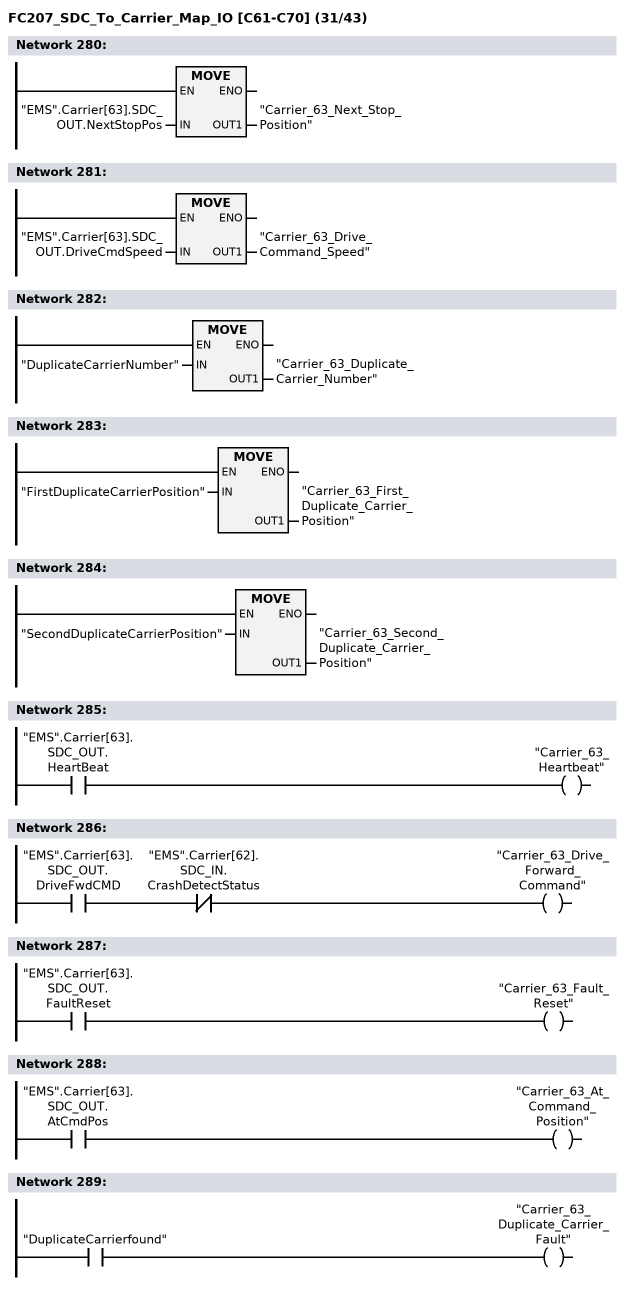
   RUNG wire#powerrail
      Move(in := "EMS".Carrier[63].SDC_OUT.NextStopPos, out1 => "Carrier_63_Next_Stop_Position")
   END_RUNG
   // the same network as SCL:
   "Carrier_63_Next_Stop_Position" := "EMS".Carrier[63].SDC_OUT.NextStopPos;
END_REGION

REGION Network 281
   RUNG wire#powerrail
      Move(in := "EMS".Carrier[63].SDC_OUT.DriveCmdSpeed, out1 => "Carrier_63_Drive_Command_Speed")
   END_RUNG
   // the same network as SCL:
   "Carrier_63_Drive_Command_Speed" := "EMS".Carrier[63].SDC_OUT.DriveCmdSpeed;
END_REGION

REGION Network 282
   RUNG wire#powerrail
      Move(in := "DuplicateCarrierNumber", out1 => "Carrier_63_Duplicate_Carrier_Number")
   END_RUNG
   // the same network as SCL:
   "Carrier_63_Duplicate_Carrier_Number" := "DuplicateCarrierNumber";
END_REGION

REGION Network 283
   RUNG wire#powerrail
      Move(in := "FirstDuplicateCarrierPosition", out1 => "Carrier_63_First_Duplicate_Carrier_Position")
   END_RUNG
   // the same network as SCL:
   "Carrier_63_First_Duplicate_Carrier_Position" := "FirstDuplicateCarrierPosition";
END_REGION

REGION Network 284
   RUNG wire#powerrail
      Move(in := "SecondDuplicateCarrierPosition", out1 => "Carrier_63_Second_Duplicate_Carrier_Position")
   END_RUNG
   // the same network as SCL:
   "Carrier_63_Second_Duplicate_Carrier_Position" := "SecondDuplicateCarrierPosition";
END_REGION

REGION Network 285
   RUNG wire#powerrail
      Contact( "EMS".Carrier[63].SDC_OUT.HeartBeat )
      Coil( "Carrier_63_Heartbeat" )
   END_RUNG
   // the same network as SCL:
   "Carrier_63_Heartbeat" := "EMS".Carrier[63].SDC_OUT.HeartBeat;
END_REGION

REGION Network 286
   RUNG wire#powerrail
      Contact( "EMS".Carrier[63].SDC_OUT.DriveFwdCMD )
      I_Contact( "EMS".Carrier[62].SDC_IN.CrashDetectStatus )
      Coil( "Carrier_63_Drive_Forward_Command" )
   END_RUNG
   // the same network as SCL:
   "Carrier_63_Drive_Forward_Command" := "EMS".Carrier[63].SDC_OUT.DriveFwdCMD AND NOT "EMS".Carrier[62].SDC_IN.CrashDetectStatus;
END_REGION

REGION Network 287
   RUNG wire#powerrail
      Contact( "EMS".Carrier[63].SDC_OUT.FaultReset )
      Coil( "Carrier_63_Fault_Reset" )
   END_RUNG
   // the same network as SCL:
   "Carrier_63_Fault_Reset" := "EMS".Carrier[63].SDC_OUT.FaultReset;
END_REGION

REGION Network 288
   RUNG wire#powerrail
      Contact( "EMS".Carrier[63].SDC_OUT.AtCmdPos )
      Coil( "Carrier_63_At_Command_Position" )
   END_RUNG
   // the same network as SCL:
   "Carrier_63_At_Command_Position" := "EMS".Carrier[63].SDC_OUT.AtCmdPos;
END_REGION

REGION Network 289
   RUNG wire#powerrail
      Contact( "DuplicateCarrierfound" )
      Coil( "Carrier_63_Duplicate_Carrier_Fault" )
   END_RUNG
   // the same network as SCL:
   "Carrier_63_Duplicate_Carrier_Fault" := "DuplicateCarrierfound";
END_REGION

REGION Network 290
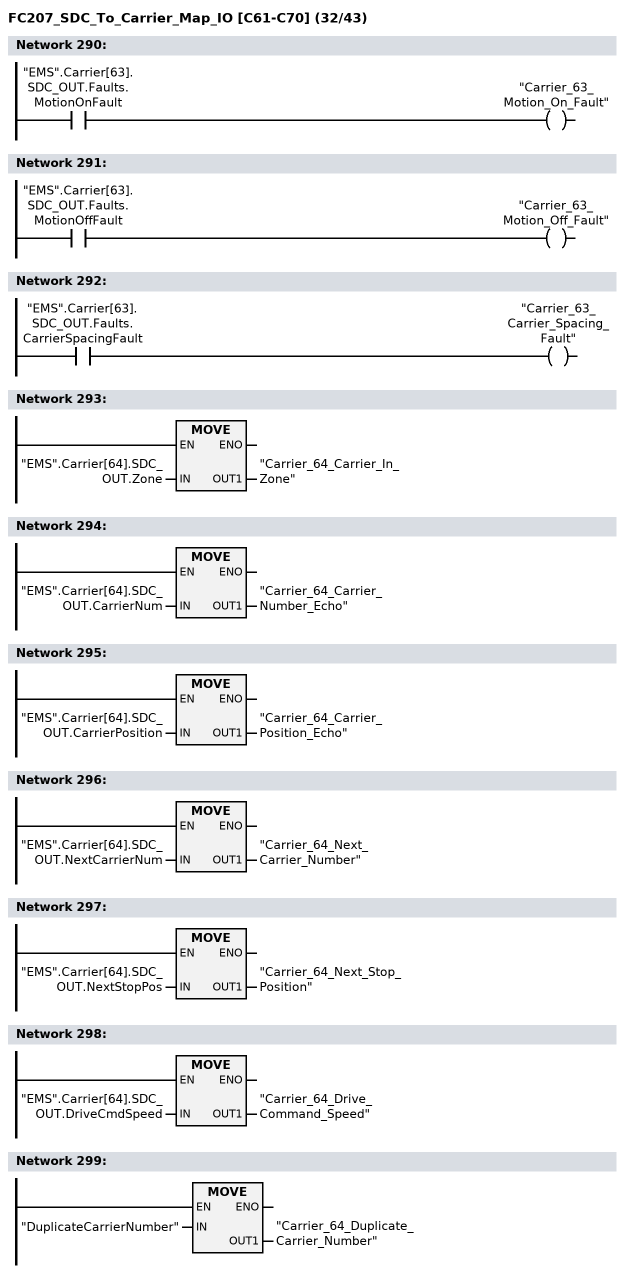
   RUNG wire#powerrail
      Contact( "EMS".Carrier[63].SDC_OUT.Faults.MotionOnFault )
      Coil( "Carrier_63_Motion_On_Fault" )
   END_RUNG
   // the same network as SCL:
   "Carrier_63_Motion_On_Fault" := "EMS".Carrier[63].SDC_OUT.Faults.MotionOnFault;
END_REGION

REGION Network 291
   RUNG wire#powerrail
      Contact( "EMS".Carrier[63].SDC_OUT.Faults.MotionOffFault )
      Coil( "Carrier_63_Motion_Off_Fault" )
   END_RUNG
   // the same network as SCL:
   "Carrier_63_Motion_Off_Fault" := "EMS".Carrier[63].SDC_OUT.Faults.MotionOffFault;
END_REGION

REGION Network 292
   RUNG wire#powerrail
      Contact( "EMS".Carrier[63].SDC_OUT.Faults.CarrierSpacingFault )
      Coil( "Carrier_63_Carrier_Spacing_Fault" )
   END_RUNG
   // the same network as SCL:
   "Carrier_63_Carrier_Spacing_Fault" := "EMS".Carrier[63].SDC_OUT.Faults.CarrierSpacingFault;
END_REGION

REGION Network 293
   RUNG wire#powerrail
      Move(in := "EMS".Carrier[64].SDC_OUT.Zone, out1 => "Carrier_64_Carrier_In_Zone")
   END_RUNG
   // the same network as SCL:
   "Carrier_64_Carrier_In_Zone" := "EMS".Carrier[64].SDC_OUT.Zone;
END_REGION

REGION Network 294
   RUNG wire#powerrail
      Move(in := "EMS".Carrier[64].SDC_OUT.CarrierNum, out1 => "Carrier_64_Carrier_Number_Echo")
   END_RUNG
   // the same network as SCL:
   "Carrier_64_Carrier_Number_Echo" := "EMS".Carrier[64].SDC_OUT.CarrierNum;
END_REGION

REGION Network 295
   RUNG wire#powerrail
      Move(in := "EMS".Carrier[64].SDC_OUT.CarrierPosition, out1 => "Carrier_64_Carrier_Position_Echo")
   END_RUNG
   // the same network as SCL:
   "Carrier_64_Carrier_Position_Echo" := "EMS".Carrier[64].SDC_OUT.CarrierPosition;
END_REGION

REGION Network 296
   RUNG wire#powerrail
      Move(in := "EMS".Carrier[64].SDC_OUT.NextCarrierNum, out1 => "Carrier_64_Next_Carrier_Number")
   END_RUNG
   // the same network as SCL:
   "Carrier_64_Next_Carrier_Number" := "EMS".Carrier[64].SDC_OUT.NextCarrierNum;
END_REGION

REGION Network 297
   RUNG wire#powerrail
      Move(in := "EMS".Carrier[64].SDC_OUT.NextStopPos, out1 => "Carrier_64_Next_Stop_Position")
   END_RUNG
   // the same network as SCL:
   "Carrier_64_Next_Stop_Position" := "EMS".Carrier[64].SDC_OUT.NextStopPos;
END_REGION

REGION Network 298
   RUNG wire#powerrail
      Move(in := "EMS".Carrier[64].SDC_OUT.DriveCmdSpeed, out1 => "Carrier_64_Drive_Command_Speed")
   END_RUNG
   // the same network as SCL:
   "Carrier_64_Drive_Command_Speed" := "EMS".Carrier[64].SDC_OUT.DriveCmdSpeed;
END_REGION

REGION Network 299
   RUNG wire#powerrail
      Move(in := "DuplicateCarrierNumber", out1 => "Carrier_64_Duplicate_Carrier_Number")
   END_RUNG
   // the same network as SCL:
   "Carrier_64_Duplicate_Carrier_Number" := "DuplicateCarrierNumber";
END_REGION

REGION Network 300
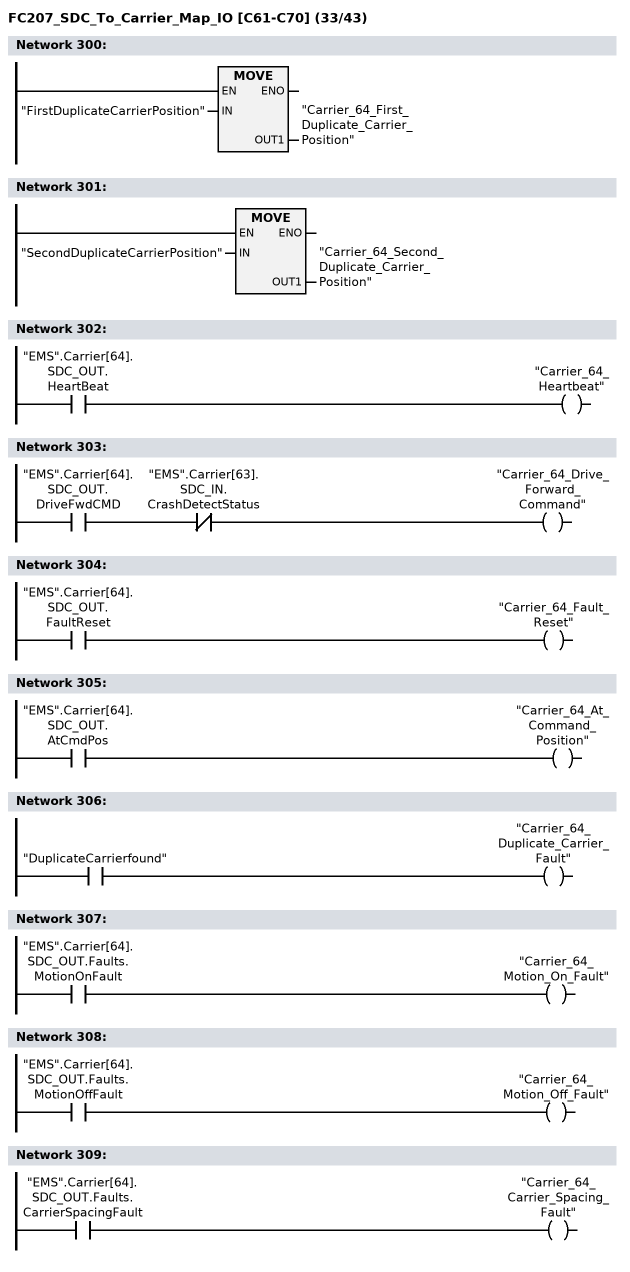
   RUNG wire#powerrail
      Move(in := "FirstDuplicateCarrierPosition", out1 => "Carrier_64_First_Duplicate_Carrier_Position")
   END_RUNG
   // the same network as SCL:
   "Carrier_64_First_Duplicate_Carrier_Position" := "FirstDuplicateCarrierPosition";
END_REGION

REGION Network 301
   RUNG wire#powerrail
      Move(in := "SecondDuplicateCarrierPosition", out1 => "Carrier_64_Second_Duplicate_Carrier_Position")
   END_RUNG
   // the same network as SCL:
   "Carrier_64_Second_Duplicate_Carrier_Position" := "SecondDuplicateCarrierPosition";
END_REGION

REGION Network 302
   RUNG wire#powerrail
      Contact( "EMS".Carrier[64].SDC_OUT.HeartBeat )
      Coil( "Carrier_64_Heartbeat" )
   END_RUNG
   // the same network as SCL:
   "Carrier_64_Heartbeat" := "EMS".Carrier[64].SDC_OUT.HeartBeat;
END_REGION

REGION Network 303
   RUNG wire#powerrail
      Contact( "EMS".Carrier[64].SDC_OUT.DriveFwdCMD )
      I_Contact( "EMS".Carrier[63].SDC_IN.CrashDetectStatus )
      Coil( "Carrier_64_Drive_Forward_Command" )
   END_RUNG
   // the same network as SCL:
   "Carrier_64_Drive_Forward_Command" := "EMS".Carrier[64].SDC_OUT.DriveFwdCMD AND NOT "EMS".Carrier[63].SDC_IN.CrashDetectStatus;
END_REGION

REGION Network 304
   RUNG wire#powerrail
      Contact( "EMS".Carrier[64].SDC_OUT.FaultReset )
      Coil( "Carrier_64_Fault_Reset" )
   END_RUNG
   // the same network as SCL:
   "Carrier_64_Fault_Reset" := "EMS".Carrier[64].SDC_OUT.FaultReset;
END_REGION

REGION Network 305
   RUNG wire#powerrail
      Contact( "EMS".Carrier[64].SDC_OUT.AtCmdPos )
      Coil( "Carrier_64_At_Command_Position" )
   END_RUNG
   // the same network as SCL:
   "Carrier_64_At_Command_Position" := "EMS".Carrier[64].SDC_OUT.AtCmdPos;
END_REGION

REGION Network 306
   RUNG wire#powerrail
      Contact( "DuplicateCarrierfound" )
      Coil( "Carrier_64_Duplicate_Carrier_Fault" )
   END_RUNG
   // the same network as SCL:
   "Carrier_64_Duplicate_Carrier_Fault" := "DuplicateCarrierfound";
END_REGION

REGION Network 307
   RUNG wire#powerrail
      Contact( "EMS".Carrier[64].SDC_OUT.Faults.MotionOnFault )
      Coil( "Carrier_64_Motion_On_Fault" )
   END_RUNG
   // the same network as SCL:
   "Carrier_64_Motion_On_Fault" := "EMS".Carrier[64].SDC_OUT.Faults.MotionOnFault;
END_REGION

REGION Network 308
   RUNG wire#powerrail
      Contact( "EMS".Carrier[64].SDC_OUT.Faults.MotionOffFault )
      Coil( "Carrier_64_Motion_Off_Fault" )
   END_RUNG
   // the same network as SCL:
   "Carrier_64_Motion_Off_Fault" := "EMS".Carrier[64].SDC_OUT.Faults.MotionOffFault;
END_REGION

REGION Network 309
   RUNG wire#powerrail
      Contact( "EMS".Carrier[64].SDC_OUT.Faults.CarrierSpacingFault )
      Coil( "Carrier_64_Carrier_Spacing_Fault" )
   END_RUNG
   // the same network as SCL:
   "Carrier_64_Carrier_Spacing_Fault" := "EMS".Carrier[64].SDC_OUT.Faults.CarrierSpacingFault;
END_REGION

REGION Network 310
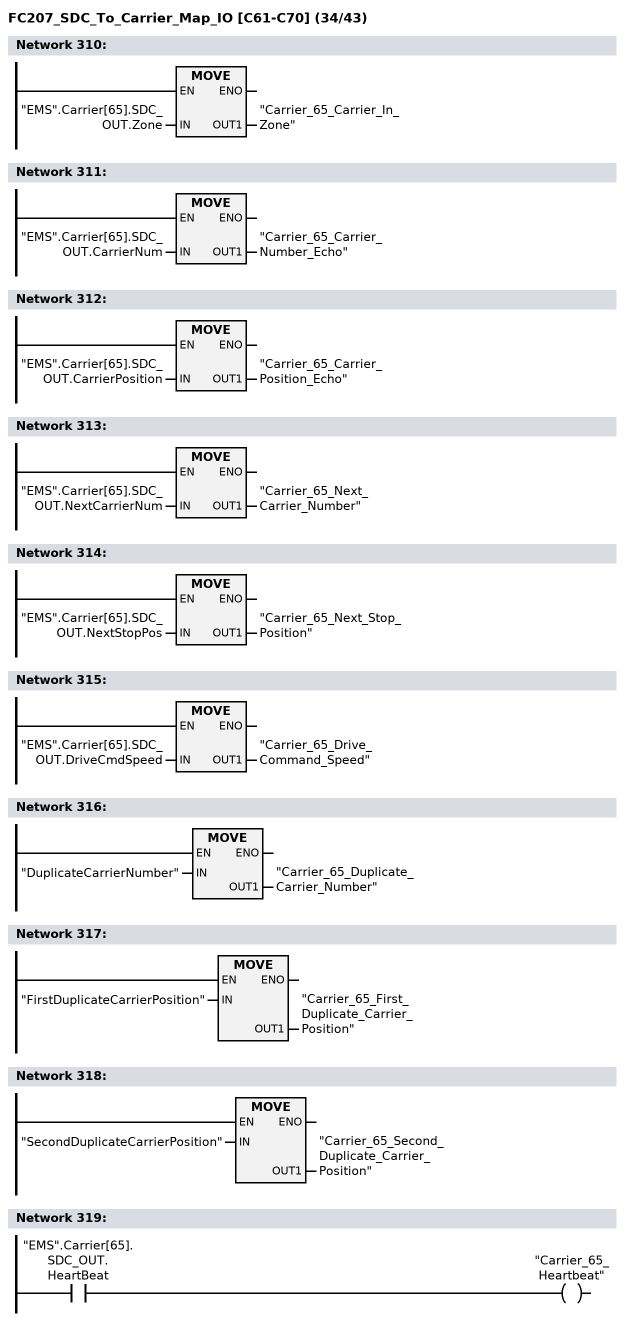
   RUNG wire#powerrail
      Move(in := "EMS".Carrier[65].SDC_OUT.Zone, out1 => "Carrier_65_Carrier_In_Zone")
   END_RUNG
   // the same network as SCL:
   "Carrier_65_Carrier_In_Zone" := "EMS".Carrier[65].SDC_OUT.Zone;
END_REGION

REGION Network 311
   RUNG wire#powerrail
      Move(in := "EMS".Carrier[65].SDC_OUT.CarrierNum, out1 => "Carrier_65_Carrier_Number_Echo")
   END_RUNG
   // the same network as SCL:
   "Carrier_65_Carrier_Number_Echo" := "EMS".Carrier[65].SDC_OUT.CarrierNum;
END_REGION

REGION Network 312
   RUNG wire#powerrail
      Move(in := "EMS".Carrier[65].SDC_OUT.CarrierPosition, out1 => "Carrier_65_Carrier_Position_Echo")
   END_RUNG
   // the same network as SCL:
   "Carrier_65_Carrier_Position_Echo" := "EMS".Carrier[65].SDC_OUT.CarrierPosition;
END_REGION

REGION Network 313
   RUNG wire#powerrail
      Move(in := "EMS".Carrier[65].SDC_OUT.NextCarrierNum, out1 => "Carrier_65_Next_Carrier_Number")
   END_RUNG
   // the same network as SCL:
   "Carrier_65_Next_Carrier_Number" := "EMS".Carrier[65].SDC_OUT.NextCarrierNum;
END_REGION

REGION Network 314
   RUNG wire#powerrail
      Move(in := "EMS".Carrier[65].SDC_OUT.NextStopPos, out1 => "Carrier_65_Next_Stop_Position")
   END_RUNG
   // the same network as SCL:
   "Carrier_65_Next_Stop_Position" := "EMS".Carrier[65].SDC_OUT.NextStopPos;
END_REGION

REGION Network 315
   RUNG wire#powerrail
      Move(in := "EMS".Carrier[65].SDC_OUT.DriveCmdSpeed, out1 => "Carrier_65_Drive_Command_Speed")
   END_RUNG
   // the same network as SCL:
   "Carrier_65_Drive_Command_Speed" := "EMS".Carrier[65].SDC_OUT.DriveCmdSpeed;
END_REGION

REGION Network 316
   RUNG wire#powerrail
      Move(in := "DuplicateCarrierNumber", out1 => "Carrier_65_Duplicate_Carrier_Number")
   END_RUNG
   // the same network as SCL:
   "Carrier_65_Duplicate_Carrier_Number" := "DuplicateCarrierNumber";
END_REGION

REGION Network 317
   RUNG wire#powerrail
      Move(in := "FirstDuplicateCarrierPosition", out1 => "Carrier_65_First_Duplicate_Carrier_Position")
   END_RUNG
   // the same network as SCL:
   "Carrier_65_First_Duplicate_Carrier_Position" := "FirstDuplicateCarrierPosition";
END_REGION

REGION Network 318
   RUNG wire#powerrail
      Move(in := "SecondDuplicateCarrierPosition", out1 => "Carrier_65_Second_Duplicate_Carrier_Position")
   END_RUNG
   // the same network as SCL:
   "Carrier_65_Second_Duplicate_Carrier_Position" := "SecondDuplicateCarrierPosition";
END_REGION

REGION Network 319
   RUNG wire#powerrail
      Contact( "EMS".Carrier[65].SDC_OUT.HeartBeat )
      Coil( "Carrier_65_Heartbeat" )
   END_RUNG
   // the same network as SCL:
   "Carrier_65_Heartbeat" := "EMS".Carrier[65].SDC_OUT.HeartBeat;
END_REGION

REGION Network 320
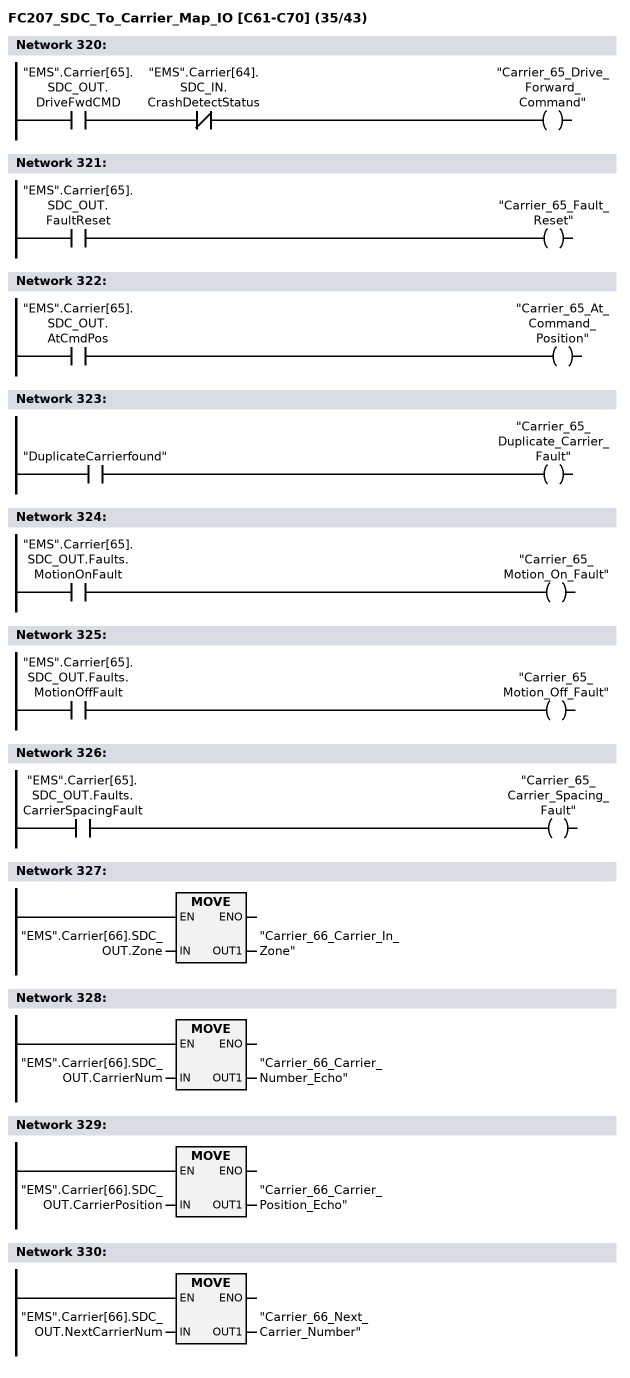
   RUNG wire#powerrail
      Contact( "EMS".Carrier[65].SDC_OUT.DriveFwdCMD )
      I_Contact( "EMS".Carrier[64].SDC_IN.CrashDetectStatus )
      Coil( "Carrier_65_Drive_Forward_Command" )
   END_RUNG
   // the same network as SCL:
   "Carrier_65_Drive_Forward_Command" := "EMS".Carrier[65].SDC_OUT.DriveFwdCMD AND NOT "EMS".Carrier[64].SDC_IN.CrashDetectStatus;
END_REGION

REGION Network 321
   RUNG wire#powerrail
      Contact( "EMS".Carrier[65].SDC_OUT.FaultReset )
      Coil( "Carrier_65_Fault_Reset" )
   END_RUNG
   // the same network as SCL:
   "Carrier_65_Fault_Reset" := "EMS".Carrier[65].SDC_OUT.FaultReset;
END_REGION

REGION Network 322
   RUNG wire#powerrail
      Contact( "EMS".Carrier[65].SDC_OUT.AtCmdPos )
      Coil( "Carrier_65_At_Command_Position" )
   END_RUNG
   // the same network as SCL:
   "Carrier_65_At_Command_Position" := "EMS".Carrier[65].SDC_OUT.AtCmdPos;
END_REGION

REGION Network 323
   RUNG wire#powerrail
      Contact( "DuplicateCarrierfound" )
      Coil( "Carrier_65_Duplicate_Carrier_Fault" )
   END_RUNG
   // the same network as SCL:
   "Carrier_65_Duplicate_Carrier_Fault" := "DuplicateCarrierfound";
END_REGION

REGION Network 324
   RUNG wire#powerrail
      Contact( "EMS".Carrier[65].SDC_OUT.Faults.MotionOnFault )
      Coil( "Carrier_65_Motion_On_Fault" )
   END_RUNG
   // the same network as SCL:
   "Carrier_65_Motion_On_Fault" := "EMS".Carrier[65].SDC_OUT.Faults.MotionOnFault;
END_REGION

REGION Network 325
   RUNG wire#powerrail
      Contact( "EMS".Carrier[65].SDC_OUT.Faults.MotionOffFault )
      Coil( "Carrier_65_Motion_Off_Fault" )
   END_RUNG
   // the same network as SCL:
   "Carrier_65_Motion_Off_Fault" := "EMS".Carrier[65].SDC_OUT.Faults.MotionOffFault;
END_REGION

REGION Network 326
   RUNG wire#powerrail
      Contact( "EMS".Carrier[65].SDC_OUT.Faults.CarrierSpacingFault )
      Coil( "Carrier_65_Carrier_Spacing_Fault" )
   END_RUNG
   // the same network as SCL:
   "Carrier_65_Carrier_Spacing_Fault" := "EMS".Carrier[65].SDC_OUT.Faults.CarrierSpacingFault;
END_REGION

REGION Network 327
   RUNG wire#powerrail
      Move(in := "EMS".Carrier[66].SDC_OUT.Zone, out1 => "Carrier_66_Carrier_In_Zone")
   END_RUNG
   // the same network as SCL:
   "Carrier_66_Carrier_In_Zone" := "EMS".Carrier[66].SDC_OUT.Zone;
END_REGION

REGION Network 328
   RUNG wire#powerrail
      Move(in := "EMS".Carrier[66].SDC_OUT.CarrierNum, out1 => "Carrier_66_Carrier_Number_Echo")
   END_RUNG
   // the same network as SCL:
   "Carrier_66_Carrier_Number_Echo" := "EMS".Carrier[66].SDC_OUT.CarrierNum;
END_REGION

REGION Network 329
   RUNG wire#powerrail
      Move(in := "EMS".Carrier[66].SDC_OUT.CarrierPosition, out1 => "Carrier_66_Carrier_Position_Echo")
   END_RUNG
   // the same network as SCL:
   "Carrier_66_Carrier_Position_Echo" := "EMS".Carrier[66].SDC_OUT.CarrierPosition;
END_REGION

REGION Network 330
   RUNG wire#powerrail
      Move(in := "EMS".Carrier[66].SDC_OUT.NextCarrierNum, out1 => "Carrier_66_Next_Carrier_Number")
   END_RUNG
   // the same network as SCL:
   "Carrier_66_Next_Carrier_Number" := "EMS".Carrier[66].SDC_OUT.NextCarrierNum;
END_REGION

REGION Network 331
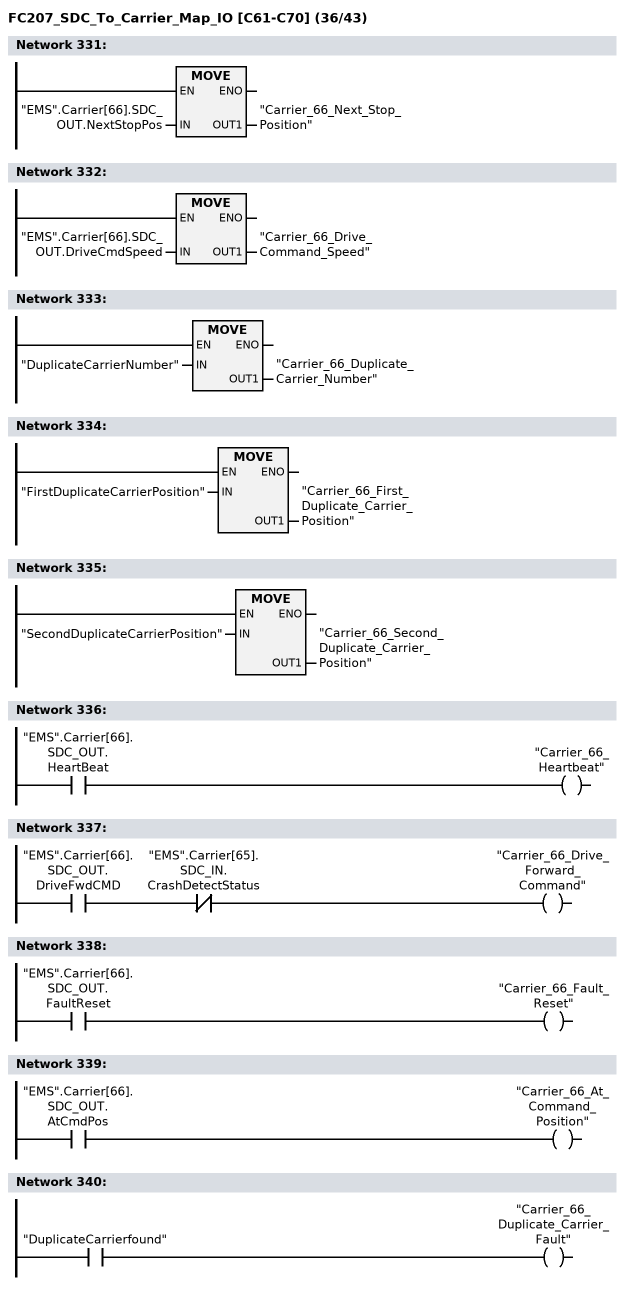
   RUNG wire#powerrail
      Move(in := "EMS".Carrier[66].SDC_OUT.NextStopPos, out1 => "Carrier_66_Next_Stop_Position")
   END_RUNG
   // the same network as SCL:
   "Carrier_66_Next_Stop_Position" := "EMS".Carrier[66].SDC_OUT.NextStopPos;
END_REGION

REGION Network 332
   RUNG wire#powerrail
      Move(in := "EMS".Carrier[66].SDC_OUT.DriveCmdSpeed, out1 => "Carrier_66_Drive_Command_Speed")
   END_RUNG
   // the same network as SCL:
   "Carrier_66_Drive_Command_Speed" := "EMS".Carrier[66].SDC_OUT.DriveCmdSpeed;
END_REGION

REGION Network 333
   RUNG wire#powerrail
      Move(in := "DuplicateCarrierNumber", out1 => "Carrier_66_Duplicate_Carrier_Number")
   END_RUNG
   // the same network as SCL:
   "Carrier_66_Duplicate_Carrier_Number" := "DuplicateCarrierNumber";
END_REGION

REGION Network 334
   RUNG wire#powerrail
      Move(in := "FirstDuplicateCarrierPosition", out1 => "Carrier_66_First_Duplicate_Carrier_Position")
   END_RUNG
   // the same network as SCL:
   "Carrier_66_First_Duplicate_Carrier_Position" := "FirstDuplicateCarrierPosition";
END_REGION

REGION Network 335
   RUNG wire#powerrail
      Move(in := "SecondDuplicateCarrierPosition", out1 => "Carrier_66_Second_Duplicate_Carrier_Position")
   END_RUNG
   // the same network as SCL:
   "Carrier_66_Second_Duplicate_Carrier_Position" := "SecondDuplicateCarrierPosition";
END_REGION

REGION Network 336
   RUNG wire#powerrail
      Contact( "EMS".Carrier[66].SDC_OUT.HeartBeat )
      Coil( "Carrier_66_Heartbeat" )
   END_RUNG
   // the same network as SCL:
   "Carrier_66_Heartbeat" := "EMS".Carrier[66].SDC_OUT.HeartBeat;
END_REGION

REGION Network 337
   RUNG wire#powerrail
      Contact( "EMS".Carrier[66].SDC_OUT.DriveFwdCMD )
      I_Contact( "EMS".Carrier[65].SDC_IN.CrashDetectStatus )
      Coil( "Carrier_66_Drive_Forward_Command" )
   END_RUNG
   // the same network as SCL:
   "Carrier_66_Drive_Forward_Command" := "EMS".Carrier[66].SDC_OUT.DriveFwdCMD AND NOT "EMS".Carrier[65].SDC_IN.CrashDetectStatus;
END_REGION

REGION Network 338
   RUNG wire#powerrail
      Contact( "EMS".Carrier[66].SDC_OUT.FaultReset )
      Coil( "Carrier_66_Fault_Reset" )
   END_RUNG
   // the same network as SCL:
   "Carrier_66_Fault_Reset" := "EMS".Carrier[66].SDC_OUT.FaultReset;
END_REGION

REGION Network 339
   RUNG wire#powerrail
      Contact( "EMS".Carrier[66].SDC_OUT.AtCmdPos )
      Coil( "Carrier_66_At_Command_Position" )
   END_RUNG
   // the same network as SCL:
   "Carrier_66_At_Command_Position" := "EMS".Carrier[66].SDC_OUT.AtCmdPos;
END_REGION

REGION Network 340
   RUNG wire#powerrail
      Contact( "DuplicateCarrierfound" )
      Coil( "Carrier_66_Duplicate_Carrier_Fault" )
   END_RUNG
   // the same network as SCL:
   "Carrier_66_Duplicate_Carrier_Fault" := "DuplicateCarrierfound";
END_REGION

REGION Network 341
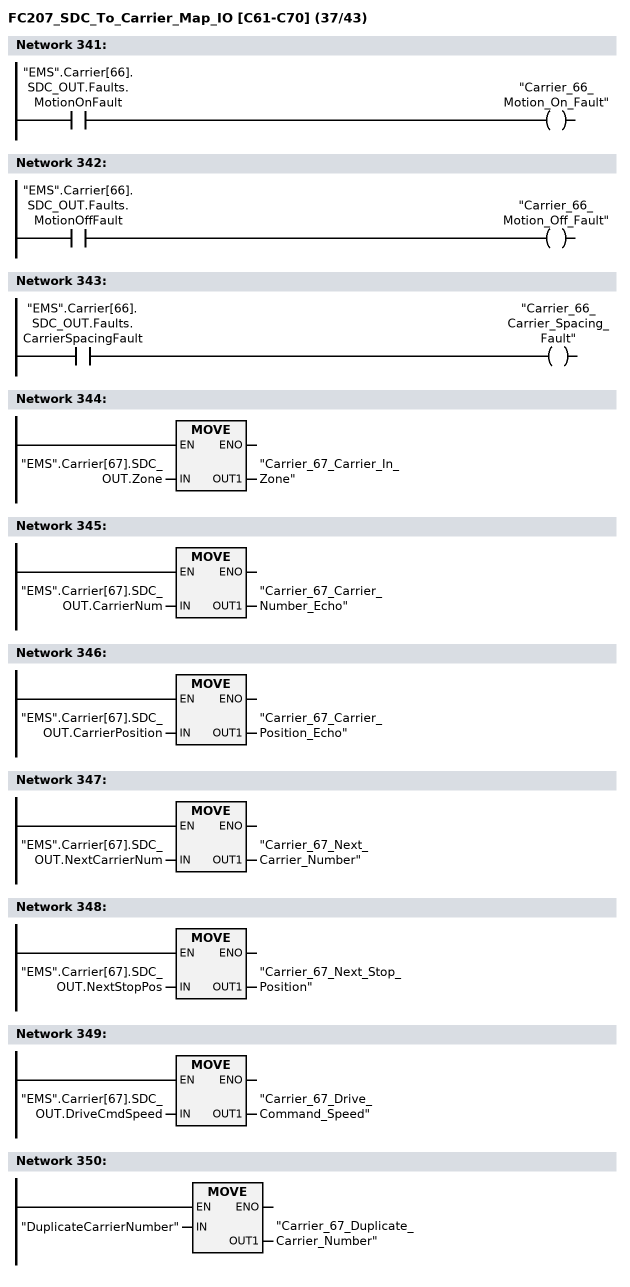
   RUNG wire#powerrail
      Contact( "EMS".Carrier[66].SDC_OUT.Faults.MotionOnFault )
      Coil( "Carrier_66_Motion_On_Fault" )
   END_RUNG
   // the same network as SCL:
   "Carrier_66_Motion_On_Fault" := "EMS".Carrier[66].SDC_OUT.Faults.MotionOnFault;
END_REGION

REGION Network 342
   RUNG wire#powerrail
      Contact( "EMS".Carrier[66].SDC_OUT.Faults.MotionOffFault )
      Coil( "Carrier_66_Motion_Off_Fault" )
   END_RUNG
   // the same network as SCL:
   "Carrier_66_Motion_Off_Fault" := "EMS".Carrier[66].SDC_OUT.Faults.MotionOffFault;
END_REGION

REGION Network 343
   RUNG wire#powerrail
      Contact( "EMS".Carrier[66].SDC_OUT.Faults.CarrierSpacingFault )
      Coil( "Carrier_66_Carrier_Spacing_Fault" )
   END_RUNG
   // the same network as SCL:
   "Carrier_66_Carrier_Spacing_Fault" := "EMS".Carrier[66].SDC_OUT.Faults.CarrierSpacingFault;
END_REGION

REGION Network 344
   RUNG wire#powerrail
      Move(in := "EMS".Carrier[67].SDC_OUT.Zone, out1 => "Carrier_67_Carrier_In_Zone")
   END_RUNG
   // the same network as SCL:
   "Carrier_67_Carrier_In_Zone" := "EMS".Carrier[67].SDC_OUT.Zone;
END_REGION

REGION Network 345
   RUNG wire#powerrail
      Move(in := "EMS".Carrier[67].SDC_OUT.CarrierNum, out1 => "Carrier_67_Carrier_Number_Echo")
   END_RUNG
   // the same network as SCL:
   "Carrier_67_Carrier_Number_Echo" := "EMS".Carrier[67].SDC_OUT.CarrierNum;
END_REGION

REGION Network 346
   RUNG wire#powerrail
      Move(in := "EMS".Carrier[67].SDC_OUT.CarrierPosition, out1 => "Carrier_67_Carrier_Position_Echo")
   END_RUNG
   // the same network as SCL:
   "Carrier_67_Carrier_Position_Echo" := "EMS".Carrier[67].SDC_OUT.CarrierPosition;
END_REGION

REGION Network 347
   RUNG wire#powerrail
      Move(in := "EMS".Carrier[67].SDC_OUT.NextCarrierNum, out1 => "Carrier_67_Next_Carrier_Number")
   END_RUNG
   // the same network as SCL:
   "Carrier_67_Next_Carrier_Number" := "EMS".Carrier[67].SDC_OUT.NextCarrierNum;
END_REGION

REGION Network 348
   RUNG wire#powerrail
      Move(in := "EMS".Carrier[67].SDC_OUT.NextStopPos, out1 => "Carrier_67_Next_Stop_Position")
   END_RUNG
   // the same network as SCL:
   "Carrier_67_Next_Stop_Position" := "EMS".Carrier[67].SDC_OUT.NextStopPos;
END_REGION

REGION Network 349
   RUNG wire#powerrail
      Move(in := "EMS".Carrier[67].SDC_OUT.DriveCmdSpeed, out1 => "Carrier_67_Drive_Command_Speed")
   END_RUNG
   // the same network as SCL:
   "Carrier_67_Drive_Command_Speed" := "EMS".Carrier[67].SDC_OUT.DriveCmdSpeed;
END_REGION

REGION Network 350
   RUNG wire#powerrail
      Move(in := "DuplicateCarrierNumber", out1 => "Carrier_67_Duplicate_Carrier_Number")
   END_RUNG
   // the same network as SCL:
   "Carrier_67_Duplicate_Carrier_Number" := "DuplicateCarrierNumber";
END_REGION

REGION Network 351
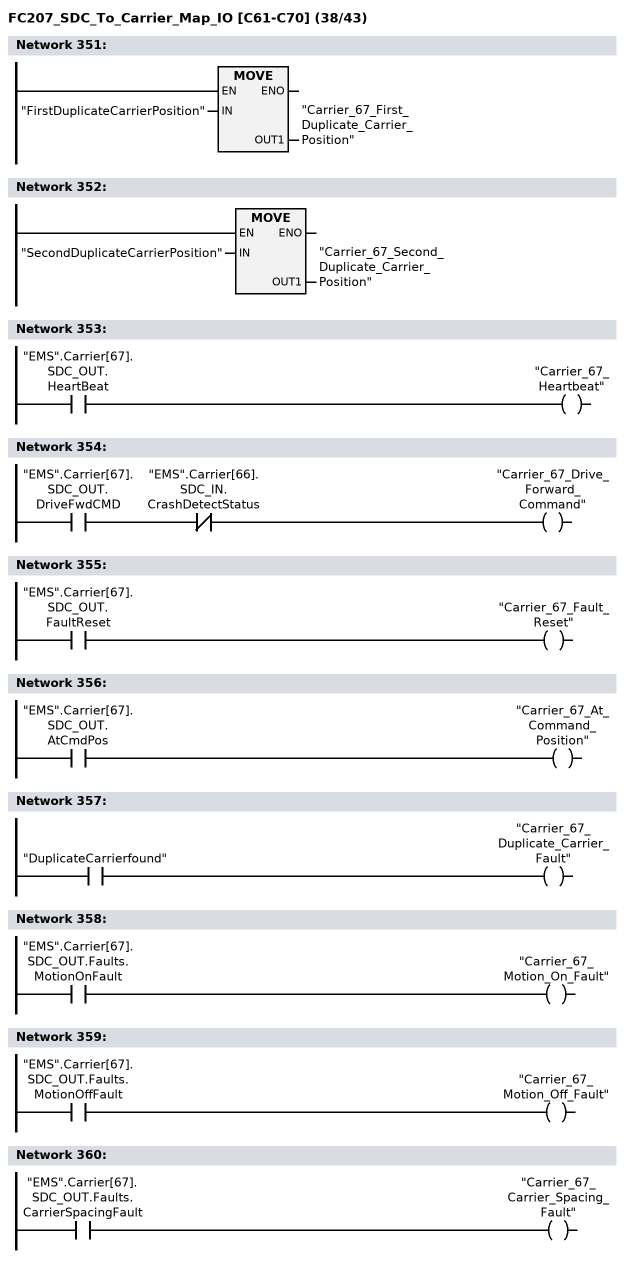
   RUNG wire#powerrail
      Move(in := "FirstDuplicateCarrierPosition", out1 => "Carrier_67_First_Duplicate_Carrier_Position")
   END_RUNG
   // the same network as SCL:
   "Carrier_67_First_Duplicate_Carrier_Position" := "FirstDuplicateCarrierPosition";
END_REGION

REGION Network 352
   RUNG wire#powerrail
      Move(in := "SecondDuplicateCarrierPosition", out1 => "Carrier_67_Second_Duplicate_Carrier_Position")
   END_RUNG
   // the same network as SCL:
   "Carrier_67_Second_Duplicate_Carrier_Position" := "SecondDuplicateCarrierPosition";
END_REGION

REGION Network 353
   RUNG wire#powerrail
      Contact( "EMS".Carrier[67].SDC_OUT.HeartBeat )
      Coil( "Carrier_67_Heartbeat" )
   END_RUNG
   // the same network as SCL:
   "Carrier_67_Heartbeat" := "EMS".Carrier[67].SDC_OUT.HeartBeat;
END_REGION

REGION Network 354
   RUNG wire#powerrail
      Contact( "EMS".Carrier[67].SDC_OUT.DriveFwdCMD )
      I_Contact( "EMS".Carrier[66].SDC_IN.CrashDetectStatus )
      Coil( "Carrier_67_Drive_Forward_Command" )
   END_RUNG
   // the same network as SCL:
   "Carrier_67_Drive_Forward_Command" := "EMS".Carrier[67].SDC_OUT.DriveFwdCMD AND NOT "EMS".Carrier[66].SDC_IN.CrashDetectStatus;
END_REGION

REGION Network 355
   RUNG wire#powerrail
      Contact( "EMS".Carrier[67].SDC_OUT.FaultReset )
      Coil( "Carrier_67_Fault_Reset" )
   END_RUNG
   // the same network as SCL:
   "Carrier_67_Fault_Reset" := "EMS".Carrier[67].SDC_OUT.FaultReset;
END_REGION

REGION Network 356
   RUNG wire#powerrail
      Contact( "EMS".Carrier[67].SDC_OUT.AtCmdPos )
      Coil( "Carrier_67_At_Command_Position" )
   END_RUNG
   // the same network as SCL:
   "Carrier_67_At_Command_Position" := "EMS".Carrier[67].SDC_OUT.AtCmdPos;
END_REGION

REGION Network 357
   RUNG wire#powerrail
      Contact( "DuplicateCarrierfound" )
      Coil( "Carrier_67_Duplicate_Carrier_Fault" )
   END_RUNG
   // the same network as SCL:
   "Carrier_67_Duplicate_Carrier_Fault" := "DuplicateCarrierfound";
END_REGION

REGION Network 358
   RUNG wire#powerrail
      Contact( "EMS".Carrier[67].SDC_OUT.Faults.MotionOnFault )
      Coil( "Carrier_67_Motion_On_Fault" )
   END_RUNG
   // the same network as SCL:
   "Carrier_67_Motion_On_Fault" := "EMS".Carrier[67].SDC_OUT.Faults.MotionOnFault;
END_REGION

REGION Network 359
   RUNG wire#powerrail
      Contact( "EMS".Carrier[67].SDC_OUT.Faults.MotionOffFault )
      Coil( "Carrier_67_Motion_Off_Fault" )
   END_RUNG
   // the same network as SCL:
   "Carrier_67_Motion_Off_Fault" := "EMS".Carrier[67].SDC_OUT.Faults.MotionOffFault;
END_REGION

REGION Network 360
   RUNG wire#powerrail
      Contact( "EMS".Carrier[67].SDC_OUT.Faults.CarrierSpacingFault )
      Coil( "Carrier_67_Carrier_Spacing_Fault" )
   END_RUNG
   // the same network as SCL:
   "Carrier_67_Carrier_Spacing_Fault" := "EMS".Carrier[67].SDC_OUT.Faults.CarrierSpacingFault;
END_REGION

REGION Network 361
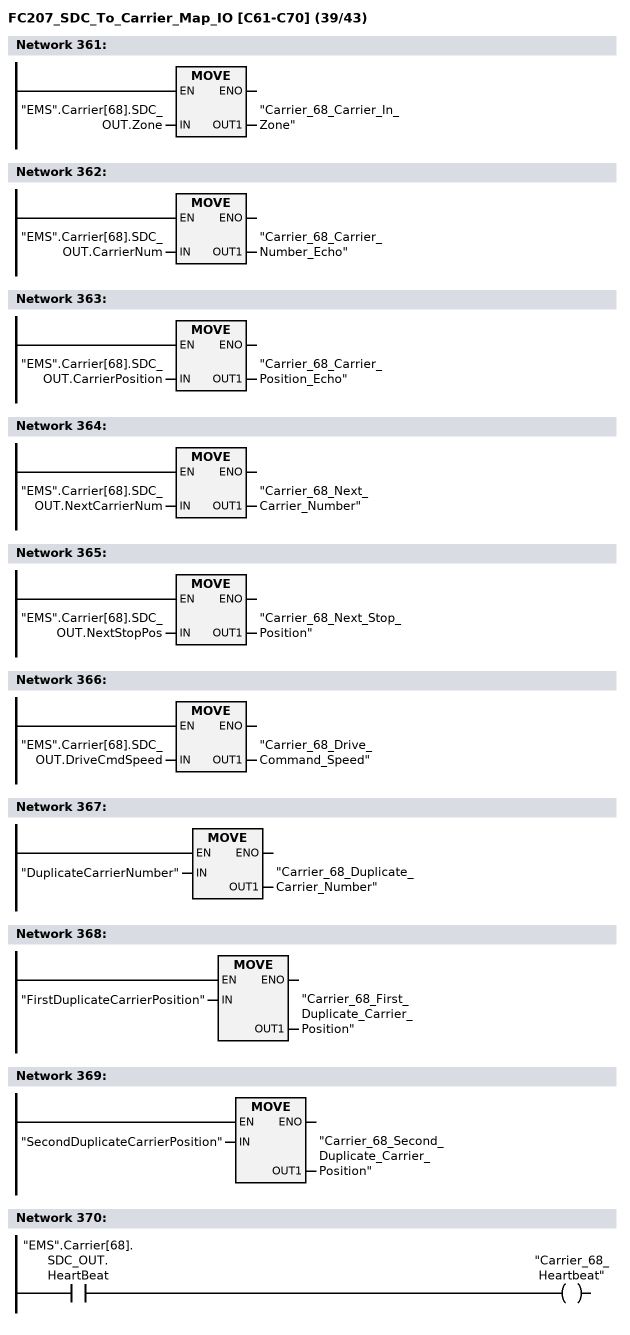
   RUNG wire#powerrail
      Move(in := "EMS".Carrier[68].SDC_OUT.Zone, out1 => "Carrier_68_Carrier_In_Zone")
   END_RUNG
   // the same network as SCL:
   "Carrier_68_Carrier_In_Zone" := "EMS".Carrier[68].SDC_OUT.Zone;
END_REGION

REGION Network 362
   RUNG wire#powerrail
      Move(in := "EMS".Carrier[68].SDC_OUT.CarrierNum, out1 => "Carrier_68_Carrier_Number_Echo")
   END_RUNG
   // the same network as SCL:
   "Carrier_68_Carrier_Number_Echo" := "EMS".Carrier[68].SDC_OUT.CarrierNum;
END_REGION

REGION Network 363
   RUNG wire#powerrail
      Move(in := "EMS".Carrier[68].SDC_OUT.CarrierPosition, out1 => "Carrier_68_Carrier_Position_Echo")
   END_RUNG
   // the same network as SCL:
   "Carrier_68_Carrier_Position_Echo" := "EMS".Carrier[68].SDC_OUT.CarrierPosition;
END_REGION
